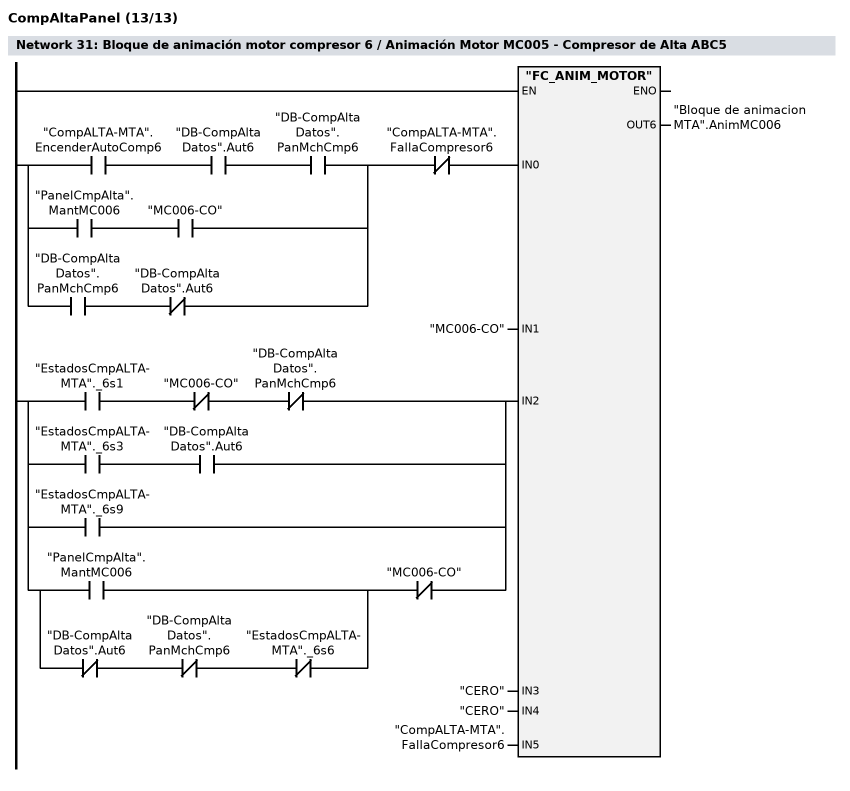
   RUNG wire#powerrail
      "FC_ANIM_MOTOR"(IN0 := wire#w2, IN2 := wire#w4, IN1 := "MC006-CO", IN3 := "CERO", IN4 := "CERO", IN5 := "CompALTA-MTA".FallaCompresor6, OUT6 => "Bloque de animacion MTA".AnimMC006)
   END_RUNG
   RUNG wire#powerrail
      Contact( "CompALTA-MTA".EncenderAutoComp6 )
      Contact( "DB-CompAltaDatos".Aut6 )
      Contact( "DB-CompAltaDatos".PanMchCmp6 )
      wire#w1
      I_Contact( "CompALTA-MTA".FallaCompresor6 )
   END_RUNG wire#w2
   RUNG wire#powerrail
      Contact( "PanelCmpAlta".MantMC006 )
      Contact( "MC006-CO" )
   END_RUNG wire#w1
   RUNG wire#powerrail
      Contact( "DB-CompAltaDatos".PanMchCmp6 )
      I_Contact( "DB-CompAltaDatos".Aut6 )
   END_RUNG wire#w1
   RUNG wire#powerrail
      Contact( "EstadosCmpALTA-MTA"._6s1 )
      I_Contact( "MC006-CO" )
      I_Contact( "DB-CompAltaDatos".PanMchCmp6 )
   END_RUNG wire#w4
   RUNG wire#powerrail
      Contact( "EstadosCmpALTA-MTA"._6s3 )
      Contact( "DB-CompAltaDatos".Aut6 )
   END_RUNG wire#w4
   RUNG wire#powerrail
      Contact( "EstadosCmpALTA-MTA"._6s9 )
   END_RUNG wire#w4
   RUNG wire#powerrail
      Contact( "PanelCmpAlta".MantMC006 )
      wire#w3
      I_Contact( "MC006-CO" )
   END_RUNG wire#w4
   RUNG wire#powerrail
      I_Contact( "DB-CompAltaDatos".Aut6 )
      I_Contact( "DB-CompAltaDatos".PanMchCmp6 )
      I_Contact( "EstadosCmpALTA-MTA"._6s6 )
   END_RUNG wire#w3
   // the same network as SCL:
   "FC_ANIM_MOTOR"(IN0 := (("CompALTA-MTA".EncenderAutoComp6 AND "DB-CompAltaDatos".Aut6 AND "DB-CompAltaDatos".PanMchCmp6) OR ("PanelCmpAlta".MantMC006 AND "MC006-CO") OR ("DB-CompAltaDatos".PanMchCmp6 AND NOT "DB-CompAltaDatos".Aut6)) AND NOT "CompALTA-MTA".FallaCompresor6,
                   IN1 := "MC006-CO",
                   IN2 := ("EstadosCmpALTA-MTA"._6s1 AND NOT "MC006-CO" AND NOT "DB-CompAltaDatos".PanMchCmp6) OR ("EstadosCmpALTA-MTA"._6s3 AND "DB-CompAltaDatos".Aut6) OR "EstadosCmpALTA-MTA"._6s9 OR (("PanelCmpAlta".MantMC006 OR (NOT "DB-CompAltaDatos".Aut6 AND NOT "DB-CompAltaDatos".PanMchCmp6 AND NOT "EstadosCmpALTA-MTA"._6s6)) AND NOT "MC006-CO"),
                   IN3 := "CERO",
                   IN4 := "CERO",
                   IN5 := "CompALTA-MTA".FallaCompresor6,
                   OUT6 => "Bloque de animacion MTA".AnimMC006);
END_REGION
END_FUNCTION

FUNCTION "ModoManualAlta" : Void   // FC48, LAD
{ S7_Optimized_Access := 'FALSE' }
VERSION : 0.1
   VAR_TEMP   // added for the SCL form of the ladder/FBD networks
      _w1 : Bool;
      _s5time1 : S5Time;
   END_VAR
BEGIN

REGION Network 1
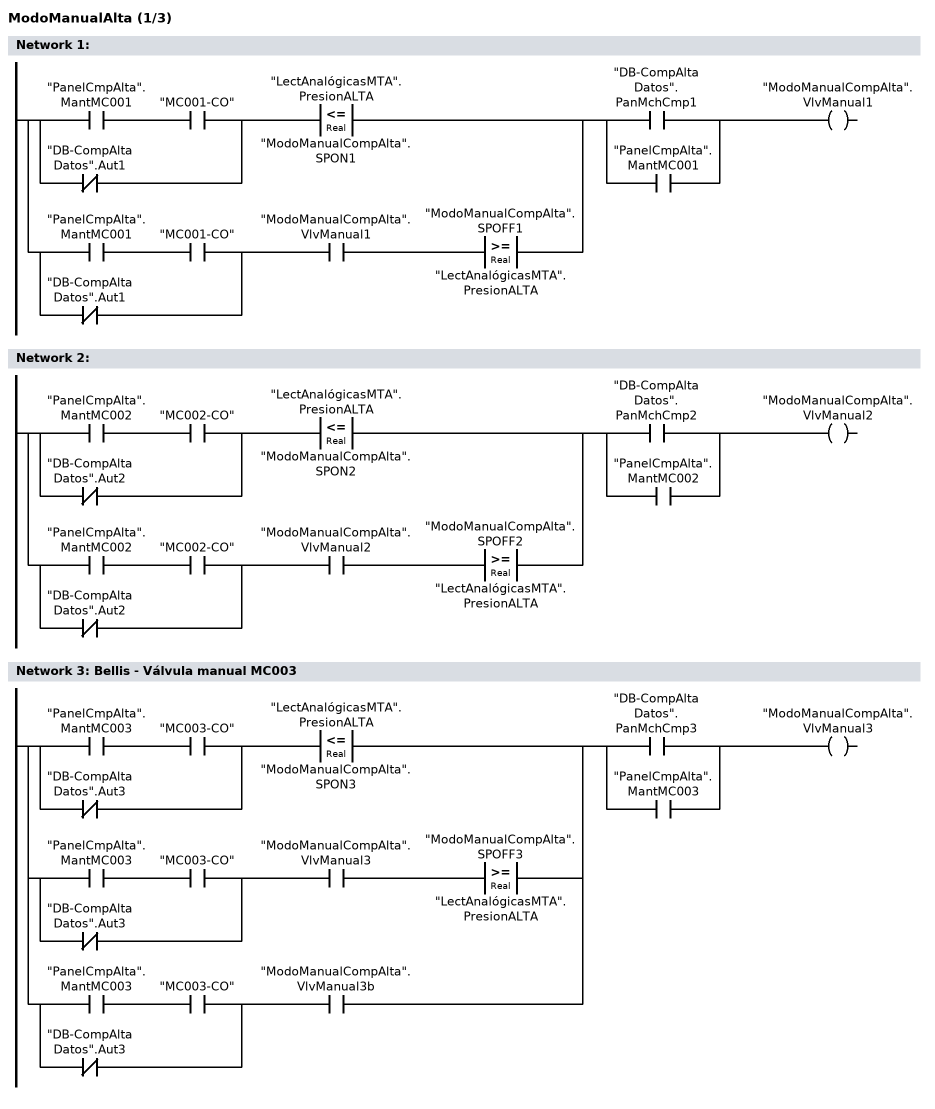
   "ModoManualCompAlta".VlvManual1 := (((NOT "DB-CompAltaDatos".Aut1 OR ("PanelCmpAlta".MantMC001 AND "MC001-CO")) AND ("LectAnalógicasMTA".PresionALTA <= "ModoManualCompAlta".SPON1)) OR ((NOT "DB-CompAltaDatos".Aut1 OR ("PanelCmpAlta".MantMC001 AND "MC001-CO")) AND "ModoManualCompAlta".VlvManual1 AND ("ModoManualCompAlta".SPOFF1 >= "LectAnalógicasMTA".PresionALTA))) AND ("DB-CompAltaDatos".PanMchCmp1 OR "PanelCmpAlta".MantMC001);
END_REGION

REGION Network 2
   "ModoManualCompAlta".VlvManual2 := (((NOT "DB-CompAltaDatos".Aut2 OR ("PanelCmpAlta".MantMC002 AND "MC002-CO")) AND ("LectAnalógicasMTA".PresionALTA <= "ModoManualCompAlta".SPON2)) OR ((NOT "DB-CompAltaDatos".Aut2 OR ("PanelCmpAlta".MantMC002 AND "MC002-CO")) AND "ModoManualCompAlta".VlvManual2 AND ("ModoManualCompAlta".SPOFF2 >= "LectAnalógicasMTA".PresionALTA))) AND ("DB-CompAltaDatos".PanMchCmp2 OR "PanelCmpAlta".MantMC002);
END_REGION

REGION Network 3: Bellis - Válvula manual MC003
   "ModoManualCompAlta".VlvManual3 := (((NOT "DB-CompAltaDatos".Aut3 OR ("PanelCmpAlta".MantMC003 AND "MC003-CO")) AND ("LectAnalógicasMTA".PresionALTA <= "ModoManualCompAlta".SPON3)) OR ((NOT "DB-CompAltaDatos".Aut3 OR ("PanelCmpAlta".MantMC003 AND "MC003-CO")) AND "ModoManualCompAlta".VlvManual3 AND ("ModoManualCompAlta".SPOFF3 >= "LectAnalógicasMTA".PresionALTA)) OR ((NOT "DB-CompAltaDatos".Aut3 OR ("PanelCmpAlta".MantMC003 AND "MC003-CO")) AND "ModoManualCompAlta".VlvManual3b)) AND ("DB-CompAltaDatos".PanMchCmp3 OR "PanelCmpAlta".MantMC003);
END_REGION

REGION Network 4: Bellis - Válvula manual MC003b
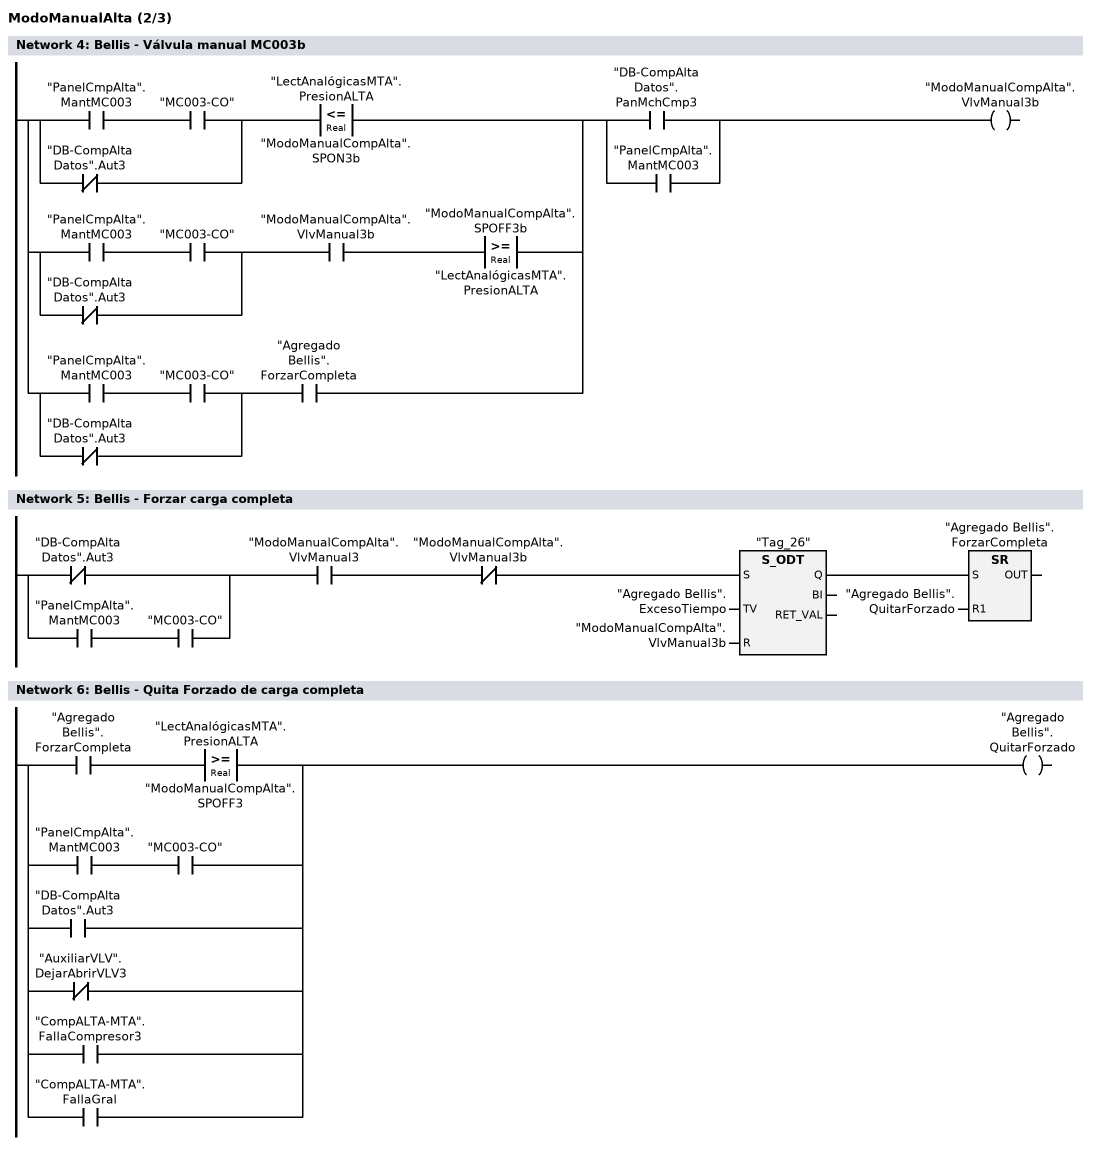
   "ModoManualCompAlta".VlvManual3b := (((NOT "DB-CompAltaDatos".Aut3 OR ("PanelCmpAlta".MantMC003 AND "MC003-CO")) AND ("LectAnalógicasMTA".PresionALTA <= "ModoManualCompAlta".SPON3b)) OR ((NOT "DB-CompAltaDatos".Aut3 OR ("PanelCmpAlta".MantMC003 AND "MC003-CO")) AND "ModoManualCompAlta".VlvManual3b AND ("ModoManualCompAlta".SPOFF3b >= "LectAnalógicasMTA".PresionALTA)) OR ((NOT "DB-CompAltaDatos".Aut3 OR ("PanelCmpAlta".MantMC003 AND "MC003-CO")) AND "Agregado Bellis".ForzarCompleta)) AND ("DB-CompAltaDatos".PanMchCmp3 OR "PanelCmpAlta".MantMC003);
END_REGION

REGION Network 5: Bellis - Forzar carga completa
   RUNG wire#powerrail
      I_Contact( "DB-CompAltaDatos".Aut3 )
      wire#w1
      Contact( "ModoManualCompAlta".VlvManual3 )
      I_Contact( "ModoManualCompAlta".VlvManual3b )
      S_ODT(T_NO := "Tag_26", TV := "Agregado Bellis".ExcesoTiempo, R := "ModoManualCompAlta".VlvManual3b, BI =>, RET_VAL =>)
      S_SR(operand := "Agregado Bellis".ForzarCompleta, r1 := "Agregado Bellis".QuitarForzado)
   END_RUNG
   RUNG wire#powerrail
      Contact( "PanelCmpAlta".MantMC003 )
      Contact( "MC003-CO" )
   END_RUNG wire#w1
   // the same network as SCL:
   #_s5time1 := S_ODT(T_NO := "Tag_26",
                      S := (NOT "DB-CompAltaDatos".Aut3 OR ("PanelCmpAlta".MantMC003 AND "MC003-CO")) AND "ModoManualCompAlta".VlvManual3 AND NOT "ModoManualCompAlta".VlvManual3b,
                      TV := "Agregado Bellis".ExcesoTiempo,
                      R := "ModoManualCompAlta".VlvManual3b,
                      Q => #_w1);
   IF #_w1 THEN
       "Agregado Bellis".ForzarCompleta := TRUE;   // SR flip-flop
   END_IF;
   IF "Agregado Bellis".QuitarForzado THEN "Agregado Bellis".ForzarCompleta := FALSE; END_IF;
END_REGION

REGION Network 6: Bellis - Quita Forzado de carga completa
   "Agregado Bellis".QuitarForzado := ("Agregado Bellis".ForzarCompleta AND ("LectAnalógicasMTA".PresionALTA >= "ModoManualCompAlta".SPOFF3)) OR "DB-CompAltaDatos".Aut3 OR ("PanelCmpAlta".MantMC003 AND "MC003-CO") OR NOT "AuxiliarVLV".DejarAbrirVLV3 OR "CompALTA-MTA".FallaCompresor3 OR "CompALTA-MTA".FallaGral;
END_REGION

REGION Network 7
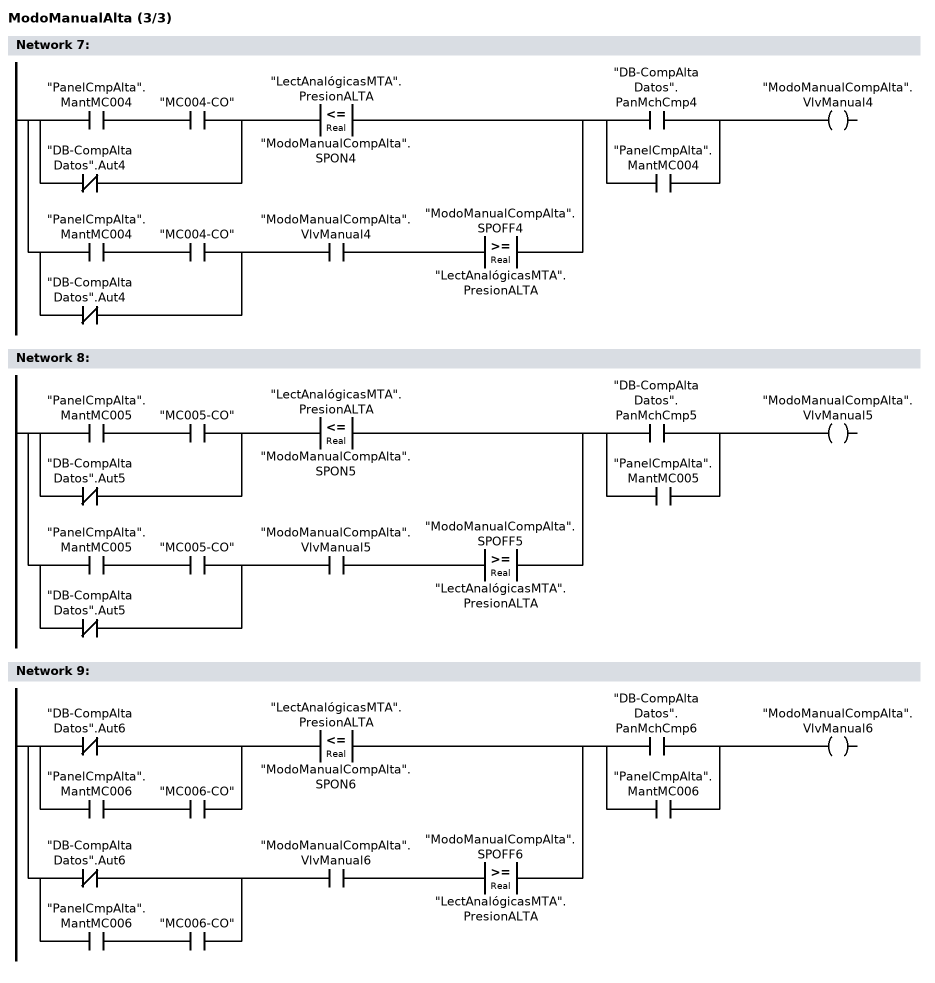
   "ModoManualCompAlta".VlvManual4 := (((NOT "DB-CompAltaDatos".Aut4 OR ("PanelCmpAlta".MantMC004 AND "MC004-CO")) AND ("LectAnalógicasMTA".PresionALTA <= "ModoManualCompAlta".SPON4)) OR ((NOT "DB-CompAltaDatos".Aut4 OR ("PanelCmpAlta".MantMC004 AND "MC004-CO")) AND "ModoManualCompAlta".VlvManual4 AND ("ModoManualCompAlta".SPOFF4 >= "LectAnalógicasMTA".PresionALTA))) AND ("DB-CompAltaDatos".PanMchCmp4 OR "PanelCmpAlta".MantMC004);
END_REGION

REGION Network 8
   "ModoManualCompAlta".VlvManual5 := (((NOT "DB-CompAltaDatos".Aut5 OR ("PanelCmpAlta".MantMC005 AND "MC005-CO")) AND ("LectAnalógicasMTA".PresionALTA <= "ModoManualCompAlta".SPON5)) OR ((NOT "DB-CompAltaDatos".Aut5 OR ("PanelCmpAlta".MantMC005 AND "MC005-CO")) AND "ModoManualCompAlta".VlvManual5 AND ("ModoManualCompAlta".SPOFF5 >= "LectAnalógicasMTA".PresionALTA))) AND ("DB-CompAltaDatos".PanMchCmp5 OR "PanelCmpAlta".MantMC005);
END_REGION

REGION Network 9
   RUNG wire#powerrail
      I_Contact( "DB-CompAltaDatos".Aut6 )
      wire#w1
      { S7_Templates := "SrcType := Real" } LE_Contact(in1 := "LectAnalógicasMTA".PresionALTA, in2 := "ModoManualCompAlta".SPON6)
      wire#w2
      Contact( "DB-CompAltaDatos".PanMchCmp6 )
      wire#w4
      Coil( "ModoManualCompAlta".VlvManual6 )
   END_RUNG
   RUNG wire#powerrail
      Contact( "PanelCmpAlta".MantMC006 )
      Contact( "MC006-CO" )
   END_RUNG wire#w1
   RUNG wire#powerrail
      I_Contact( "DB-CompAltaDatos".Aut6 )
      wire#w3
      Contact( "ModoManualCompAlta".VlvManual6 )
      { S7_Templates := "SrcType := Real" } GE_Contact(in1 := "ModoManualCompAlta".SPOFF6, in2 := "LectAnalógicasMTA".PresionALTA)
   END_RUNG wire#w2
   RUNG wire#powerrail
      Contact( "PanelCmpAlta".MantMC006 )
      Contact( "MC006-CO" )
   END_RUNG wire#w3
   RUNG wire#w2
      Contact( "PanelCmpAlta".MantMC006 )
   END_RUNG wire#w4
   // the same network as SCL:
   "ModoManualCompAlta".VlvManual6 := (((NOT "DB-CompAltaDatos".Aut6 OR ("PanelCmpAlta".MantMC006 AND "MC006-CO")) AND ("LectAnalógicasMTA".PresionALTA <= "ModoManualCompAlta".SPON6)) OR ((NOT "DB-CompAltaDatos".Aut6 OR ("PanelCmpAlta".MantMC006 AND "MC006-CO")) AND "ModoManualCompAlta".VlvManual6 AND ("ModoManualCompAlta".SPOFF6 >= "LectAnalógicasMTA".PresionALTA))) AND ("DB-CompAltaDatos".PanMchCmp6 OR "PanelCmpAlta".MantMC006);
END_REGION
END_FUNCTION

FUNCTION "PurgaComAlta" : Void   // FC51, LAD
{ S7_Optimized_Access := 'FALSE' }
VERSION : 0.1
// Control de electrovalvulas para realizar purga de compresores, evitando simultaneidad. Con habilitación y seteos de tiempos desde panel.
   VAR_TEMP   // added for the SCL form of the ladder/FBD networks
      _w1 : Bool;
      _s5time1 : S5Time;
      _s5time2 : S5Time;
   END_VAR
BEGIN

REGION Network 1
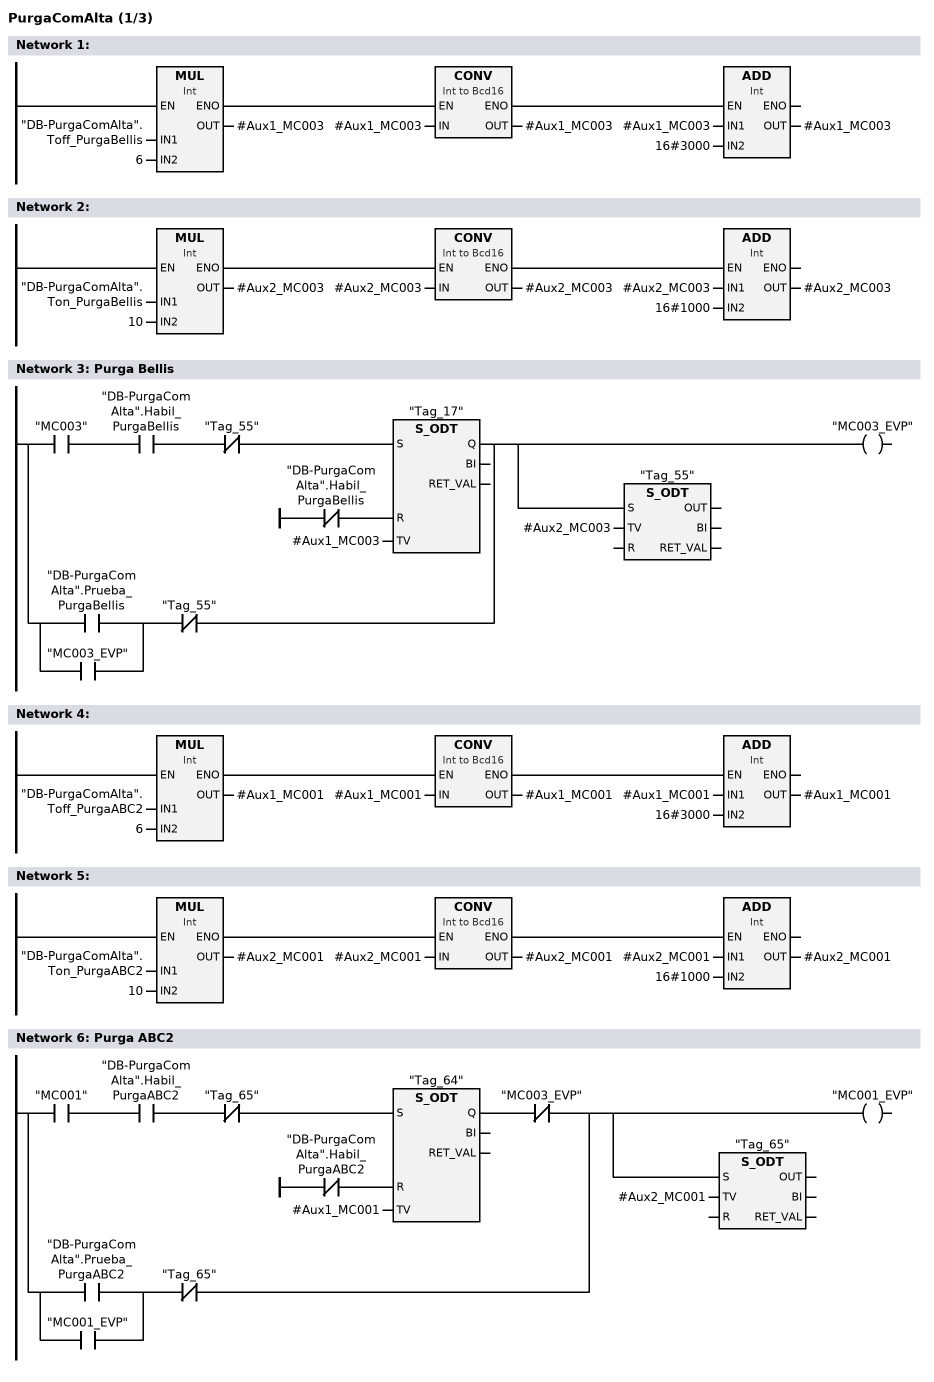
   RUNG wire#powerrail
      { S7_Templates := "SrcType := Int"; S7_GenerateENO := "TRUE" } Mul(in1 := "DB-PurgaComAlta".Toff_PurgaBellis, in2 := 6, out => #Aux1_MC003)
      { S7_Templates := "[SrcType := Int, DestType := Bcd16]"; S7_GenerateENO := "TRUE" } Convert(in := #Aux1_MC003, out => #Aux1_MC003)
      { S7_Templates := "SrcType := Int"; S7_GenerateENO := "TRUE" } Add(in1 := #Aux1_MC003, in2 := 16#3000, out => #Aux1_MC003)
   END_RUNG
   // the same network as SCL:
   // ENO of a box is taken as its EN; it also drops when the box reports an error
   #Aux1_MC003 := "DB-PurgaComAlta".Toff_PurgaBellis * 6;
   #Aux1_MC003 := INT_TO_BCD16(#Aux1_MC003);
   #Aux1_MC003 := #Aux1_MC003 + 16#3000;
END_REGION

REGION Network 2
   RUNG wire#powerrail
      { S7_Templates := "SrcType := Int"; S7_GenerateENO := "TRUE" } Mul(in1 := "DB-PurgaComAlta".Ton_PurgaBellis, in2 := 10, out => #Aux2_MC003)
      { S7_Templates := "[SrcType := Int, DestType := Bcd16]"; S7_GenerateENO := "TRUE" } Convert(in := #Aux2_MC003, out => #Aux2_MC003)
      { S7_Templates := "SrcType := Int"; S7_GenerateENO := "TRUE" } Add(in1 := #Aux2_MC003, in2 := 16#1000, out => #Aux2_MC003)
   END_RUNG
   // the same network as SCL:
   // ENO of a box is taken as its EN; it also drops when the box reports an error
   #Aux2_MC003 := "DB-PurgaComAlta".Ton_PurgaBellis * 10;
   #Aux2_MC003 := INT_TO_BCD16(#Aux2_MC003);
   #Aux2_MC003 := #Aux2_MC003 + 16#1000;
END_REGION

REGION Network 3: Purga Bellis
   RUNG wire#powerrail
      Contact( "MC003" )
      Contact( "DB-PurgaComAlta".Habil_PurgaBellis )
      I_Contact( "Tag_55" )
      S_ODT(T_NO := "Tag_17", R := wire#w1, TV := #Aux1_MC003, BI =>, RET_VAL =>)
      wire#w2
      Coil( "MC003_EVP" )
   END_RUNG
   RUNG wire#powerrail
      I_Contact( "DB-PurgaComAlta".Habil_PurgaBellis )
   END_RUNG wire#w1
   RUNG wire#powerrail
      Contact( "DB-PurgaComAlta".Prueba_PurgaBellis )
      wire#w3
      I_Contact( "Tag_55" )
   END_RUNG wire#w2
   RUNG wire#powerrail
      Contact( "MC003_EVP" )
   END_RUNG wire#w3
   RUNG wire#w2
      S_ODT(T_NO := "Tag_55", TV := #Aux2_MC003, R :=, BI =>, RET_VAL =>)
   END_RUNG
   // the same network as SCL:
   #_s5time1 := S_ODT(T_NO := "Tag_17",
                      S := "MC003" AND "DB-PurgaComAlta".Habil_PurgaBellis AND NOT "Tag_55",
                      R := NOT "DB-PurgaComAlta".Habil_PurgaBellis,
                      TV := #Aux1_MC003,
                      Q => #_w1);
   "MC003_EVP" := #_w1 OR (("DB-PurgaComAlta".Prueba_PurgaBellis OR "MC003_EVP") AND NOT "Tag_55");
   #_s5time2 := S_ODT(T_NO := "Tag_55", S := "MC003_EVP", TV := #Aux2_MC003);
END_REGION

REGION Network 4
   RUNG wire#powerrail
      { S7_Templates := "SrcType := Int"; S7_GenerateENO := "TRUE" } Mul(in1 := "DB-PurgaComAlta".Toff_PurgaABC2, in2 := 6, out => #Aux1_MC001)
      { S7_Templates := "[SrcType := Int, DestType := Bcd16]"; S7_GenerateENO := "TRUE" } Convert(in := #Aux1_MC001, out => #Aux1_MC001)
      { S7_Templates := "SrcType := Int"; S7_GenerateENO := "TRUE" } Add(in1 := #Aux1_MC001, in2 := 16#3000, out => #Aux1_MC001)
   END_RUNG
   // the same network as SCL:
   // ENO of a box is taken as its EN; it also drops when the box reports an error
   #Aux1_MC001 := "DB-PurgaComAlta".Toff_PurgaABC2 * 6;
   #Aux1_MC001 := INT_TO_BCD16(#Aux1_MC001);
   #Aux1_MC001 := #Aux1_MC001 + 16#3000;
END_REGION

REGION Network 5
   RUNG wire#powerrail
      { S7_Templates := "SrcType := Int"; S7_GenerateENO := "TRUE" } Mul(in1 := "DB-PurgaComAlta".Ton_PurgaABC2, in2 := 10, out => #Aux2_MC001)
      { S7_Templates := "[SrcType := Int, DestType := Bcd16]"; S7_GenerateENO := "TRUE" } Convert(in := #Aux2_MC001, out => #Aux2_MC001)
      { S7_Templates := "SrcType := Int"; S7_GenerateENO := "TRUE" } Add(in1 := #Aux2_MC001, in2 := 16#1000, out => #Aux2_MC001)
   END_RUNG
   // the same network as SCL:
   // ENO of a box is taken as its EN; it also drops when the box reports an error
   #Aux2_MC001 := "DB-PurgaComAlta".Ton_PurgaABC2 * 10;
   #Aux2_MC001 := INT_TO_BCD16(#Aux2_MC001);
   #Aux2_MC001 := #Aux2_MC001 + 16#1000;
END_REGION

REGION Network 6: Purga ABC2
   RUNG wire#powerrail
      Contact( "MC001" )
      Contact( "DB-PurgaComAlta".Habil_PurgaABC2 )
      I_Contact( "Tag_65" )
      S_ODT(T_NO := "Tag_64", R := wire#w1, TV := #Aux1_MC001, BI =>, RET_VAL =>)
      I_Contact( "MC003_EVP" )
      wire#w2
      Coil( "MC001_EVP" )
   END_RUNG
   RUNG wire#powerrail
      I_Contact( "DB-PurgaComAlta".Habil_PurgaABC2 )
   END_RUNG wire#w1
   RUNG wire#powerrail
      Contact( "DB-PurgaComAlta".Prueba_PurgaABC2 )
      wire#w3
      I_Contact( "Tag_65" )
   END_RUNG wire#w2
   RUNG wire#powerrail
      Contact( "MC001_EVP" )
   END_RUNG wire#w3
   RUNG wire#w2
      S_ODT(T_NO := "Tag_65", TV := #Aux2_MC001, R :=, BI =>, RET_VAL =>)
   END_RUNG
   // the same network as SCL:
   #_s5time1 := S_ODT(T_NO := "Tag_64",
                      S := "MC001" AND "DB-PurgaComAlta".Habil_PurgaABC2 AND NOT "Tag_65",
                      R := NOT "DB-PurgaComAlta".Habil_PurgaABC2,
                      TV := #Aux1_MC001,
                      Q => #_w1);
   "MC001_EVP" := (#_w1 AND NOT "MC003_EVP") OR (("DB-PurgaComAlta".Prueba_PurgaABC2 OR "MC001_EVP") AND NOT "Tag_65");
   #_s5time2 := S_ODT(T_NO := "Tag_65", S := "MC001_EVP", TV := #Aux2_MC001);
END_REGION

REGION Network 7
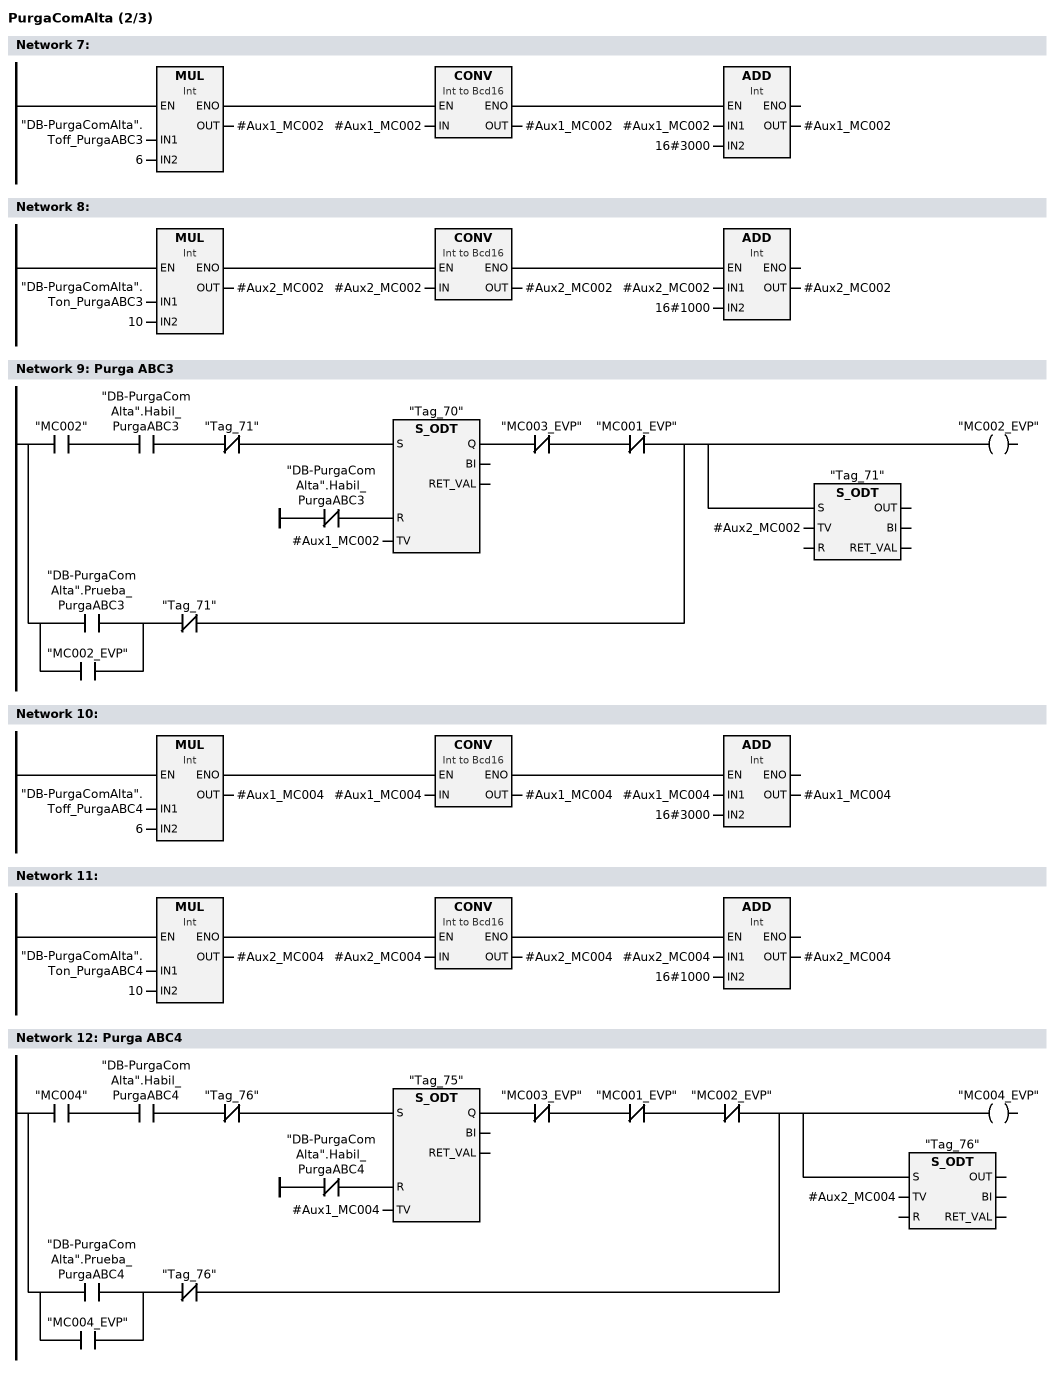
   RUNG wire#powerrail
      { S7_Templates := "SrcType := Int"; S7_GenerateENO := "TRUE" } Mul(in1 := "DB-PurgaComAlta".Toff_PurgaABC3, in2 := 6, out => #Aux1_MC002)
      { S7_Templates := "[SrcType := Int, DestType := Bcd16]"; S7_GenerateENO := "TRUE" } Convert(in := #Aux1_MC002, out => #Aux1_MC002)
      { S7_Templates := "SrcType := Int"; S7_GenerateENO := "TRUE" } Add(in1 := #Aux1_MC002, in2 := 16#3000, out => #Aux1_MC002)
   END_RUNG
   // the same network as SCL:
   // ENO of a box is taken as its EN; it also drops when the box reports an error
   #Aux1_MC002 := "DB-PurgaComAlta".Toff_PurgaABC3 * 6;
   #Aux1_MC002 := INT_TO_BCD16(#Aux1_MC002);
   #Aux1_MC002 := #Aux1_MC002 + 16#3000;
END_REGION

REGION Network 8
   RUNG wire#powerrail
      { S7_Templates := "SrcType := Int"; S7_GenerateENO := "TRUE" } Mul(in1 := "DB-PurgaComAlta".Ton_PurgaABC3, in2 := 10, out => #Aux2_MC002)
      { S7_Templates := "[SrcType := Int, DestType := Bcd16]"; S7_GenerateENO := "TRUE" } Convert(in := #Aux2_MC002, out => #Aux2_MC002)
      { S7_Templates := "SrcType := Int"; S7_GenerateENO := "TRUE" } Add(in1 := #Aux2_MC002, in2 := 16#1000, out => #Aux2_MC002)
   END_RUNG
   // the same network as SCL:
   // ENO of a box is taken as its EN; it also drops when the box reports an error
   #Aux2_MC002 := "DB-PurgaComAlta".Ton_PurgaABC3 * 10;
   #Aux2_MC002 := INT_TO_BCD16(#Aux2_MC002);
   #Aux2_MC002 := #Aux2_MC002 + 16#1000;
END_REGION

REGION Network 9: Purga ABC3
   RUNG wire#powerrail
      Contact( "MC002" )
      Contact( "DB-PurgaComAlta".Habil_PurgaABC3 )
      I_Contact( "Tag_71" )
      S_ODT(T_NO := "Tag_70", R := wire#w1, TV := #Aux1_MC002, BI =>, RET_VAL =>)
      I_Contact( "MC003_EVP" )
      I_Contact( "MC001_EVP" )
      wire#w2
      Coil( "MC002_EVP" )
   END_RUNG
   RUNG wire#powerrail
      I_Contact( "DB-PurgaComAlta".Habil_PurgaABC3 )
   END_RUNG wire#w1
   RUNG wire#powerrail
      Contact( "DB-PurgaComAlta".Prueba_PurgaABC3 )
      wire#w3
      I_Contact( "Tag_71" )
   END_RUNG wire#w2
   RUNG wire#powerrail
      Contact( "MC002_EVP" )
   END_RUNG wire#w3
   RUNG wire#w2
      S_ODT(T_NO := "Tag_71", TV := #Aux2_MC002, R :=, BI =>, RET_VAL =>)
   END_RUNG
   // the same network as SCL:
   #_s5time1 := S_ODT(T_NO := "Tag_70",
                      S := "MC002" AND "DB-PurgaComAlta".Habil_PurgaABC3 AND NOT "Tag_71",
                      R := NOT "DB-PurgaComAlta".Habil_PurgaABC3,
                      TV := #Aux1_MC002,
                      Q => #_w1);
   "MC002_EVP" := (#_w1 AND NOT "MC003_EVP" AND NOT "MC001_EVP") OR (("DB-PurgaComAlta".Prueba_PurgaABC3 OR "MC002_EVP") AND NOT "Tag_71");
   #_s5time2 := S_ODT(T_NO := "Tag_71", S := "MC002_EVP", TV := #Aux2_MC002);
END_REGION

REGION Network 10
   RUNG wire#powerrail
      { S7_Templates := "SrcType := Int"; S7_GenerateENO := "TRUE" } Mul(in1 := "DB-PurgaComAlta".Toff_PurgaABC4, in2 := 6, out => #Aux1_MC004)
      { S7_Templates := "[SrcType := Int, DestType := Bcd16]"; S7_GenerateENO := "TRUE" } Convert(in := #Aux1_MC004, out => #Aux1_MC004)
      { S7_Templates := "SrcType := Int"; S7_GenerateENO := "TRUE" } Add(in1 := #Aux1_MC004, in2 := 16#3000, out => #Aux1_MC004)
   END_RUNG
   // the same network as SCL:
   // ENO of a box is taken as its EN; it also drops when the box reports an error
   #Aux1_MC004 := "DB-PurgaComAlta".Toff_PurgaABC4 * 6;
   #Aux1_MC004 := INT_TO_BCD16(#Aux1_MC004);
   #Aux1_MC004 := #Aux1_MC004 + 16#3000;
END_REGION

REGION Network 11
   RUNG wire#powerrail
      { S7_Templates := "SrcType := Int"; S7_GenerateENO := "TRUE" } Mul(in1 := "DB-PurgaComAlta".Ton_PurgaABC4, in2 := 10, out => #Aux2_MC004)
      { S7_Templates := "[SrcType := Int, DestType := Bcd16]"; S7_GenerateENO := "TRUE" } Convert(in := #Aux2_MC004, out => #Aux2_MC004)
      { S7_Templates := "SrcType := Int"; S7_GenerateENO := "TRUE" } Add(in1 := #Aux2_MC004, in2 := 16#1000, out => #Aux2_MC004)
   END_RUNG
   // the same network as SCL:
   // ENO of a box is taken as its EN; it also drops when the box reports an error
   #Aux2_MC004 := "DB-PurgaComAlta".Ton_PurgaABC4 * 10;
   #Aux2_MC004 := INT_TO_BCD16(#Aux2_MC004);
   #Aux2_MC004 := #Aux2_MC004 + 16#1000;
END_REGION

REGION Network 12: Purga ABC4
   RUNG wire#powerrail
      Contact( "MC004" )
      Contact( "DB-PurgaComAlta".Habil_PurgaABC4 )
      I_Contact( "Tag_76" )
      S_ODT(T_NO := "Tag_75", R := wire#w1, TV := #Aux1_MC004, BI =>, RET_VAL =>)
      I_Contact( "MC003_EVP" )
      I_Contact( "MC001_EVP" )
      I_Contact( "MC002_EVP" )
      wire#w2
      Coil( "MC004_EVP" )
   END_RUNG
   RUNG wire#powerrail
      I_Contact( "DB-PurgaComAlta".Habil_PurgaABC4 )
   END_RUNG wire#w1
   RUNG wire#powerrail
      Contact( "DB-PurgaComAlta".Prueba_PurgaABC4 )
      wire#w3
      I_Contact( "Tag_76" )
   END_RUNG wire#w2
   RUNG wire#powerrail
      Contact( "MC004_EVP" )
   END_RUNG wire#w3
   RUNG wire#w2
      S_ODT(T_NO := "Tag_76", TV := #Aux2_MC004, R :=, BI =>, RET_VAL =>)
   END_RUNG
   // the same network as SCL:
   #_s5time1 := S_ODT(T_NO := "Tag_75",
                      S := "MC004" AND "DB-PurgaComAlta".Habil_PurgaABC4 AND NOT "Tag_76",
                      R := NOT "DB-PurgaComAlta".Habil_PurgaABC4,
                      TV := #Aux1_MC004,
                      Q => #_w1);
   "MC004_EVP" := (#_w1 AND NOT "MC003_EVP" AND NOT "MC001_EVP" AND NOT "MC002_EVP") OR (("DB-PurgaComAlta".Prueba_PurgaABC4 OR "MC004_EVP") AND NOT "Tag_76");
   #_s5time2 := S_ODT(T_NO := "Tag_76", S := "MC004_EVP", TV := #Aux2_MC004);
END_REGION

REGION Network 13
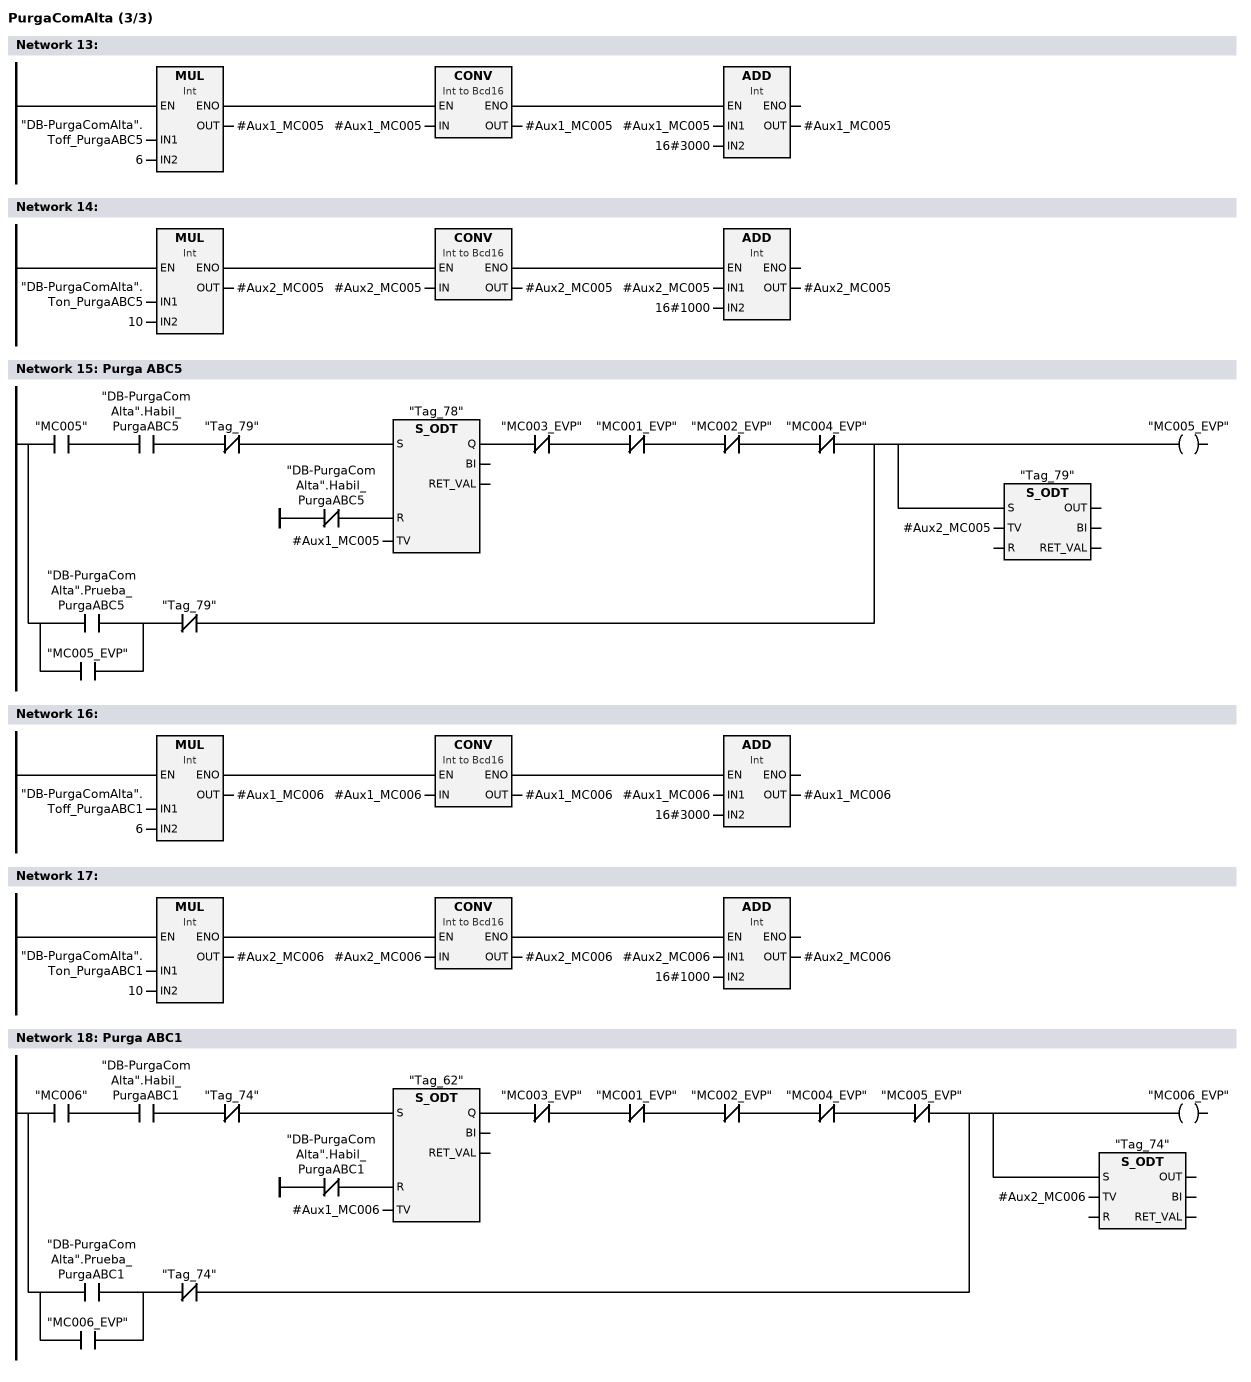
   RUNG wire#powerrail
      { S7_Templates := "SrcType := Int"; S7_GenerateENO := "TRUE" } Mul(in1 := "DB-PurgaComAlta".Toff_PurgaABC5, in2 := 6, out => #Aux1_MC005)
      { S7_Templates := "[SrcType := Int, DestType := Bcd16]"; S7_GenerateENO := "TRUE" } Convert(in := #Aux1_MC005, out => #Aux1_MC005)
      { S7_Templates := "SrcType := Int"; S7_GenerateENO := "TRUE" } Add(in1 := #Aux1_MC005, in2 := 16#3000, out => #Aux1_MC005)
   END_RUNG
   // the same network as SCL:
   // ENO of a box is taken as its EN; it also drops when the box reports an error
   #Aux1_MC005 := "DB-PurgaComAlta".Toff_PurgaABC5 * 6;
   #Aux1_MC005 := INT_TO_BCD16(#Aux1_MC005);
   #Aux1_MC005 := #Aux1_MC005 + 16#3000;
END_REGION

REGION Network 14
   RUNG wire#powerrail
      { S7_Templates := "SrcType := Int"; S7_GenerateENO := "TRUE" } Mul(in1 := "DB-PurgaComAlta".Ton_PurgaABC5, in2 := 10, out => #Aux2_MC005)
      { S7_Templates := "[SrcType := Int, DestType := Bcd16]"; S7_GenerateENO := "TRUE" } Convert(in := #Aux2_MC005, out => #Aux2_MC005)
      { S7_Templates := "SrcType := Int"; S7_GenerateENO := "TRUE" } Add(in1 := #Aux2_MC005, in2 := 16#1000, out => #Aux2_MC005)
   END_RUNG
   // the same network as SCL:
   // ENO of a box is taken as its EN; it also drops when the box reports an error
   #Aux2_MC005 := "DB-PurgaComAlta".Ton_PurgaABC5 * 10;
   #Aux2_MC005 := INT_TO_BCD16(#Aux2_MC005);
   #Aux2_MC005 := #Aux2_MC005 + 16#1000;
END_REGION

REGION Network 15: Purga ABC5
   RUNG wire#powerrail
      Contact( "MC005" )
      Contact( "DB-PurgaComAlta".Habil_PurgaABC5 )
      I_Contact( "Tag_79" )
      S_ODT(T_NO := "Tag_78", R := wire#w1, TV := #Aux1_MC005, BI =>, RET_VAL =>)
      I_Contact( "MC003_EVP" )
      I_Contact( "MC001_EVP" )
      I_Contact( "MC002_EVP" )
      I_Contact( "MC004_EVP" )
      wire#w2
      Coil( "MC005_EVP" )
   END_RUNG
   RUNG wire#powerrail
      I_Contact( "DB-PurgaComAlta".Habil_PurgaABC5 )
   END_RUNG wire#w1
   RUNG wire#powerrail
      Contact( "DB-PurgaComAlta".Prueba_PurgaABC5 )
      wire#w3
      I_Contact( "Tag_79" )
   END_RUNG wire#w2
   RUNG wire#powerrail
      Contact( "MC005_EVP" )
   END_RUNG wire#w3
   RUNG wire#w2
      S_ODT(T_NO := "Tag_79", TV := #Aux2_MC005, R :=, BI =>, RET_VAL =>)
   END_RUNG
   // the same network as SCL:
   #_s5time1 := S_ODT(T_NO := "Tag_78",
                      S := "MC005" AND "DB-PurgaComAlta".Habil_PurgaABC5 AND NOT "Tag_79",
                      R := NOT "DB-PurgaComAlta".Habil_PurgaABC5,
                      TV := #Aux1_MC005,
                      Q => #_w1);
   "MC005_EVP" := (#_w1 AND NOT "MC003_EVP" AND NOT "MC001_EVP" AND NOT "MC002_EVP" AND NOT "MC004_EVP") OR (("DB-PurgaComAlta".Prueba_PurgaABC5 OR "MC005_EVP") AND NOT "Tag_79");
   #_s5time2 := S_ODT(T_NO := "Tag_79", S := "MC005_EVP", TV := #Aux2_MC005);
END_REGION

REGION Network 16
   RUNG wire#powerrail
      { S7_Templates := "SrcType := Int"; S7_GenerateENO := "TRUE" } Mul(in1 := "DB-PurgaComAlta".Toff_PurgaABC1, in2 := 6, out => #Aux1_MC006)
      { S7_Templates := "[SrcType := Int, DestType := Bcd16]"; S7_GenerateENO := "TRUE" } Convert(in := #Aux1_MC006, out => #Aux1_MC006)
      { S7_Templates := "SrcType := Int"; S7_GenerateENO := "TRUE" } Add(in1 := #Aux1_MC006, in2 := 16#3000, out => #Aux1_MC006)
   END_RUNG
   // the same network as SCL:
   // ENO of a box is taken as its EN; it also drops when the box reports an error
   #Aux1_MC006 := "DB-PurgaComAlta".Toff_PurgaABC1 * 6;
   #Aux1_MC006 := INT_TO_BCD16(#Aux1_MC006);
   #Aux1_MC006 := #Aux1_MC006 + 16#3000;
END_REGION

REGION Network 17
   RUNG wire#powerrail
      { S7_Templates := "SrcType := Int"; S7_GenerateENO := "TRUE" } Mul(in1 := "DB-PurgaComAlta".Ton_PurgaABC1, in2 := 10, out => #Aux2_MC006)
      { S7_Templates := "[SrcType := Int, DestType := Bcd16]"; S7_GenerateENO := "TRUE" } Convert(in := #Aux2_MC006, out => #Aux2_MC006)
      { S7_Templates := "SrcType := Int"; S7_GenerateENO := "TRUE" } Add(in1 := #Aux2_MC006, in2 := 16#1000, out => #Aux2_MC006)
   END_RUNG
   // the same network as SCL:
   // ENO of a box is taken as its EN; it also drops when the box reports an error
   #Aux2_MC006 := "DB-PurgaComAlta".Ton_PurgaABC1 * 10;
   #Aux2_MC006 := INT_TO_BCD16(#Aux2_MC006);
   #Aux2_MC006 := #Aux2_MC006 + 16#1000;
END_REGION
